// TIA Portal project "Praca_Przejsciowa_S7-1200" (V15.1)
// Vorlageprojekt für das Buch mit Zielsystem S7-1200

(* hardware
DEVICE "S7-1200-Station_1"  S7-1200 Station
   slot 0: "Baugruppenträger_0"  Rack  V1.0
   slot 1: "PLC_1"  CPU 1211C DC/DC/DC  6ES7 211-1AE40-0XB0  V4.1
DEVICE "PC-System_1"  SIMATIC PC station
   slot 0: "SIMATIC PC station"  Rail  SIMATIC PC-Station  V1.0
      slot 125: "Stationmanager"  Station_Manager  V6.0.4
   slot 1: "HMI_RT_1"  WinCC RT Advanced  6AV2 104-0xxxx-xxxx  15.1.0.0
      slot 33792: "Host interface"  Host interface
   slot 2: "IE general_1"  IE General  IE_CP  V8.2.0
*)

// ===== PLC "PLC_1"  CPU 1211C DC/DC/DC =====

VAR_GLOBAL   // PLC tag table "Standard-Variablentabelle"
   "Tag_1" AT %A0.0 : Bool;
   "Tag_2" AT %E0.0 : Bool;
   "Tag_3" AT %E0.1 : Bool;
   "Tag_4" AT %ID30 : DWord;
   "Tag_5" AT %IW32 : Word;
   "Tag_6" AT %IW36 : Int;
   "Tag_7" AT %IW40 : Int;
   "Tag_8" AT %IW30 : Int;
   "Tag_9" AT %IW3 : Word;
   "Tag_10" AT %IW34 : Int;
   "Tag_11" AT %QW30 : Int;
   "Tag_12" AT %QW32 : Int;
   "Tag_13" AT %QW34 : Int;
   "Tag_14" AT %QW40 : Int;
   "Tag_15" AT %QW42 : Int;
   "Tag_16" AT %QW44 : Int;
   "Tag_17" AT %IW38 : Int;
   "Discharge1" AT %MW10 : Int;
   "ALARM_WORD" AT %MW0 : Word;
END_VAR

// folder: DBs

DATA_BLOCK "ExchangeData"   // DB1
{ S7_Optimized_Access := 'FALSE' }
VERSION : 0.1
   VAR
      iT1_LVL : Int;   // Poziom wody w zbiorniku 1
      iT1_DIS_FL : Int;   // Przepływ na wylocie zbiornika 1
      iT1_SP : Int := 150;   // Wartość zadana regulacji w zbiorniku 1
      rT1_MV : Real;   // Wartość sterowania dla zbiornika 1
      rT1_H_REG : Real := 10.0;   // Szerokość strefy histerezy regulatora zbiornika 1
      rT1_B_REG : Real := 100.0;   // Wzmocnienie przekaźnika (Zbiornik 1)
      xT1_HH_ALM : Bool;   // Alarm poziomu HH Zbiornik 1
      xT1_H_ALM : Bool;   // Alarm poziomu H Zbiornik 1
      xT1_L_ALM : Bool;   // Alarm poziomu L Zbiornik 1
      xT1_LL_ALM : Bool;   // Alarm poziomu LL Zbiornik 1
      xT1_VLV_ALM : Bool;   // Alarm – awaria zaworu Zbiornik 1
      iT2_LVL : Int;   // Poziom wody w zbiorniku 2
      iT2_DIS_FL : Int;   // Przepływ na wylocie zbiornika 2
      iT2_SP : Int := 150;   // Wartość zadana regulacji w zbiorniku 2
      rT2_MV : Real;   // Wartość sterowania dla zbiornika 2
      rT2_P_REG : Real := 5.0;   // Wzmocnienie regulatora Zbiornik 2
      rT2_I_REG : Real := 5.0;   // Parametr I regulatora Zbiornik 2
      rT2_D_REG : Real;   // Parametr D regulatora Zbiornik 2
      xT2_HH_ALM : Bool;   // Alarm poziomu HH Zbiornik 2
      xT2_H_ALM : Bool;   // Alarm poziomu H Zbiornik 2
      xT2_L_ALM : Bool;   // Alarm poziomu L Zbiornik 2
      xT2_LL_ALM : Bool;   // Alarm poziomu LL Zbiornik 2
      xT2_VLV_ALM : Bool;   // Alarm – awaria zaworu Zbiornik 2
      iT3_LVL : Int;   // Poziom wody w zbiorniku 3
      iT3_DIS_FL : Int;   // Przepływ na wylocie zbiornika 3
      iT3_SP : Int := 150;   // Wartość zadana regulacji w zbiorniku 3
      rT3_MV : Real;   // Wartość sterowania dla zbiornika 3
      rT3_P_REG : Real := 5.0;   // Wzmocnienie regulatora Zbiornik 3
      rT3_I_REG : Real := 10.0;   // Parametr I regulatora Zbiornik 3
      rT3_B_REG : Real := 100.0;   // Wzmocnienie przekaźnika Zbiornik 3
      xT3_HH_ALM : Bool;   // Alarm poziomu HH Zbiornik 3
      xT3_H_ALM : Bool;   // Alarm poziomu H Zbiornik 3
      xT3_L_ALM : Bool;   // Alarm poziomu L Zbiornik 3
      xT3_LL_ALM : Bool;   // Alarm poziomu LL Zbiornik 3
      xT3_VLV_ALM : Bool;   // Alarm – awaria zaworu Zbiornik 3
   END_VAR
BEGIN
END_DATA_BLOCK

DATA_BLOCK "Tank1 Control_DB"   // DB4
{ S7_Optimized_Access := 'TRUE' }
VERSION : 0.1
// stored: InstanceOfName Tank1 Control
"Tank1 Control"
BEGIN
END_DATA_BLOCK

DATA_BLOCK "Disturbance Generator_DB"   // DB5
{ S7_Optimized_Access := 'TRUE' }
VERSION : 0.1
// stored: InstanceOfName Disturbance Generator
"Disturbance Generator"
BEGIN
END_DATA_BLOCK

DATA_BLOCK "Tank 2 Control_DB"   // DB8
{ S7_Optimized_Access := 'TRUE' }
VERSION : 0.1
// stored: InstanceOfName Tank 2 Control
"Tank 2 Control"
BEGIN
END_DATA_BLOCK

DATA_BLOCK "Tank 3 Control_DB"   // DB9
{ S7_Optimized_Access := 'TRUE' }
VERSION : 0.1
// stored: InstanceOfName Tank 3 Control
"Tank 3 Control"
BEGIN
END_DATA_BLOCK

// folder: IO

DATA_BLOCK "Input_DB"   // DB2
{ S7_Optimized_Access := 'TRUE' }
VERSION : 0.1
// stored: InstanceOfName Input
"Input"
BEGIN
END_DATA_BLOCK

DATA_BLOCK "Output_DB"   // DB3
{ S7_Optimized_Access := 'TRUE' }
VERSION : 0.1
// stored: InstanceOfName Output
"Output"
BEGIN
END_DATA_BLOCK

// folder: (top level)

FUNCTION_BLOCK "Tank1 Control"   // FB3, LAD
{ S7_Optimized_Access := 'TRUE' }
VERSION : 0.1
   VAR_INPUT
      Level : Int;
      SP : Int := 150;
      h_reg : Real := 10.0;
      B_reg : Real := 100.0;
      HH_LVL : Int := 280;
      H_LVL : Int := 250;
      L_LVL : Int := 50;
      LL_LVL : Int := 20;
   END_VAR
   VAR_OUTPUT
      HH_Alarm : Bool;
      H_Alarm : Bool;
      L_Alarm : Bool;
      LL_Alarm : Bool;
      Vlv_Pos_Alarm : Bool;
      MV : Real;
   END_VAR
   VAR
      prev_control : Bool;
      control_action : Bool;
   END_VAR
BEGIN

REGION Network 1 (SCL)
   REGION Level control

       IF #Level < #SP - #h_reg THEN
           #control_action := 1;
       ELSIF #Level > #SP + #h_reg THEN
           #control_action := 0;
       ELSE
           #control_action := #prev_control;
       END_IF;

       #prev_control := #control_action;

       #MV := BOOL_TO_INT(#control_action) * #B_reg;


   END_REGION


   REGION ALARMS
       #HH_Alarm := FALSE;
       #H_Alarm := FALSE;
       #LL_Alarm := FALSE;
       #L_Alarm := FALSE;

       IF #Level > #HH_LVL THEN
           #HH_Alarm := TRUE;
       ELSIF #Level > #H_LVL THEN
           #H_Alarm := TRUE;
       END_IF;

       IF #Level < #LL_LVL THEN
           #LL_Alarm := TRUE;
       ELSIF #Level < #L_LVL THEN
           #L_Alarm := TRUE;
       END_IF;

   END_REGION
END_REGION
END_FUNCTION_BLOCK

FUNCTION_BLOCK "Disturbance Generator"   // FB4, LAD
{ S7_Optimized_Access := 'TRUE' }
VERSION : 0.1
   VAR_INPUT
      minOpen : Int;
      maxOpen : Int := 100;
   END_VAR
   VAR_OUTPUT
      iT1_Dis_vlv : Int;
      iT2_Dis_vlv : Int;
      iT3_Dis_vlv : Int;
   END_VAR
   VAR
      rDistrbance_T1 : Real := 50.0;
      rDistrbance_T2 : Real := 50.0;
      rDistrbance_T3 : Real := 50.0;
      rDisturbanceDesire : Real := 40.0;
      xDistrubanceRising : Bool;
   END_VAR
   VAR_TEMP
      temp_time : DTL;
      Seed1 : Real;
      Seed2 : Real;
      dist1 : Real;
      dist2 : Real;
      dist3 : Real;
   END_VAR
BEGIN

REGION Network 1 (SCL)
   // Symulacja zmian otwarcia zaworu na wyjściu jako zakłócenia
   // Seed generation from system clock
   #Seed1 := RD_SYS_T(#temp_time);
   #Seed1 := #temp_time.SECOND;
   #Seed2 := #temp_time.NANOSECOND;
   //fast and randomly changing distrubance
   #dist1 := SIN(#Seed1) + SIN(#Seed2);
   #dist1 := COS(#Seed1) + SIN(#Seed2);
   #dist1 := COS(#Seed1) + COS(#Seed2);

   // Slowly changing opennig between 20-70%
   IF #xDistrubanceRising THEN
       #rDisturbanceDesire := #rDisturbanceDesire + 0.05;
   ELSE
       #rDisturbanceDesire := #rDisturbanceDesire - 0.05;
   END_IF;

   IF #rDisturbanceDesire < 20.0 THEN
       #xDistrubanceRising := TRUE;
   ELSIF #rDisturbanceDesire > 70.0 THEN
       #xDistrubanceRising := FALSE;
   END_IF;

   // Position is sum of random distrubance and factor pushing it to
   // slowly changing desired position
   #rDistrbance_T1 := #rDistrbance_T1 + 0.1 * #dist1 + 0.01*(#rDisturbanceDesire - #rDistrbance_T1);
   #rDistrbance_T2 := #rDistrbance_T2 + 0.1 * #dist2 + 0.01 * (#rDisturbanceDesire - #rDistrbance_T2);
   #rDistrbance_T3 := #rDistrbance_T3 + 0.1 * #dist3 + 0.01 * (#rDisturbanceDesire - #rDistrbance_T3);

   // Position limited between 5-95%
   #iT1_Dis_vlv := LIMIT(MN := 5, IN := #rDistrbance_T1, MX := 95);
   #iT2_Dis_vlv := LIMIT(MN := 5, IN := #rDistrbance_T2, MX := 95);
   #iT3_Dis_vlv := LIMIT(MN := 5, IN := #rDistrbance_T3, MX := 95);
END_REGION
END_FUNCTION_BLOCK

FUNCTION_BLOCK "Tank 2 Control"   // FB5, SCL
{ S7_Optimized_Access := 'TRUE' }
VERSION : 0.1
   VAR_INPUT
      Level : Int := 0;
      SP : Int := 150;
      P_reg : Real := 10.0;
      I_reg : Real := 10.0;
      HH_LVL : Int := 280;
      H_LVL : Int := 250;
      L_LVL : Int := 50;
      LL_LVL : Int := 20;
   END_VAR
   VAR_OUTPUT
      HH_Alarm : Bool := false;
      H_Alarm : Bool := false;
      L_Alarm : Bool := false;
      LL_Alarm : Bool := false;
      Vlv_Pos_Alarm : Bool := false;
      MV : Real := 0.0;
   END_VAR
   VAR
      I_action : Real := 0.0;
      Error : Real;
      Executed : Bool;
   END_VAR
   VAR_TEMP
      P_action : Real;
   END_VAR
   VAR CONSTANT
      Interval : Time := T#100ms;
      rInterval_ms : Real := 100.0;
   END_VAR
BEGIN
   // PID opration handled by OB30
   // for constant interval time

   REGION ALARMS
       #HH_Alarm := FALSE;
       #H_Alarm := FALSE;
       #LL_Alarm := FALSE;
       #L_Alarm := FALSE;

       IF #Level > #HH_LVL THEN
           #HH_Alarm := TRUE;
       ELSIF #Level > #H_LVL THEN
           #H_Alarm := TRUE;
       END_IF;

       IF #Level < #LL_LVL THEN
           #LL_Alarm := TRUE;
       ELSIF #Level < #L_LVL THEN
           #L_Alarm := TRUE;
       END_IF;

   END_REGION
END_FUNCTION_BLOCK

FUNCTION_BLOCK "Tank 3 Control"   // FB6, LAD
{ S7_Optimized_Access := 'TRUE' }
VERSION : 0.1
   VAR_INPUT
      Level : Int;
      SP : Int := 150;
      P_reg : Real := 5.0;
      I_reg : Real := 10.0;
      B_reg : Real := 100.0;
      HH_LVL : Int := 280;
      H_LVL : Int := 250;
      L_LVL : Int := 50;
      LL_LVL : Int := 20;
   END_VAR
   VAR_OUTPUT
      HH_Alarm : Bool := false;
      H_Alarm : Bool := false;
      L_Alarm : Bool := false;
      LL_Alarm : Bool := false;
      Vlv_Pos_Alarm : Bool := false;
      MV : Real := 0.0;
   END_VAR
   VAR
      I_action : Real := 0.0;
      Error : Real := 0.0;
      Ref_sig : Real := 0.0;
      Control_sig : Real := 0.0;
      Ref_sig_period : Real := 5.0;   // okres sygnały piłokształtnego
   END_VAR
BEGIN

REGION Network 1
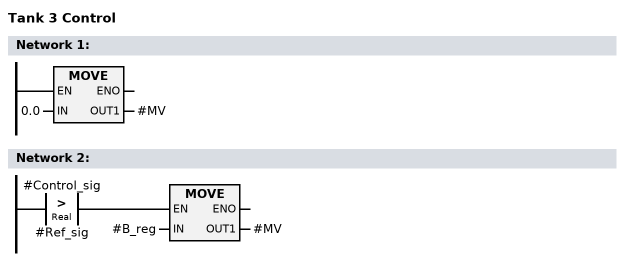
   RUNG wire#powerrail
      Move(in := 0.0, out1 => #MV)
   END_RUNG
   // the same network as SCL:
   #MV := 0.0;
END_REGION

REGION Network 2
   RUNG wire#powerrail
      { S7_Templates := "SrcType := Real" } GT_Contact(in1 := #Control_sig, in2 := #Ref_sig)
      Move(in := #B_reg, out1 => #MV)
   END_RUNG
   // the same network as SCL:
   IF #Control_sig > #Ref_sig THEN #MV := #B_reg; END_IF;
END_REGION

REGION Network 3 (SCL)
   // PID opration handled by OB31
   // for constant interval time

   REGION ALARMS
       #HH_Alarm := FALSE;
       #H_Alarm := FALSE;
       #LL_Alarm := FALSE;
       #L_Alarm := FALSE;

       IF #Level > #HH_LVL THEN
           #HH_Alarm := TRUE;
       ELSIF #Level > #H_LVL THEN
           #H_Alarm := TRUE;
       END_IF;

       IF #Level < #LL_LVL THEN
           #LL_Alarm := TRUE;
       ELSIF #Level < #L_LVL THEN
           #L_Alarm := TRUE;
       END_IF;

   END_REGION
END_REGION
END_FUNCTION_BLOCK

ORGANIZATION_BLOCK "Main"   // OB1, LAD, ProgramCycle
TITLE = "Main Program Sweep (Cycle)"
{ S7_Optimized_Access := 'TRUE' }
VERSION : 0.1
   VAR_INPUT
      Initial_Call : Bool;   // Initial call of this OB
      Remanence : Bool;   // =True, if remanent data are available
   END_VAR
BEGIN

REGION Network 1: Konnektierungsbaustein für PLC-Lab
   // Im Netzwerk 1 wird der Konnektierungsbaustein für PLC-Lab aufgerufen.
   // Dieser Aufruf darf nicht entfernt werden!
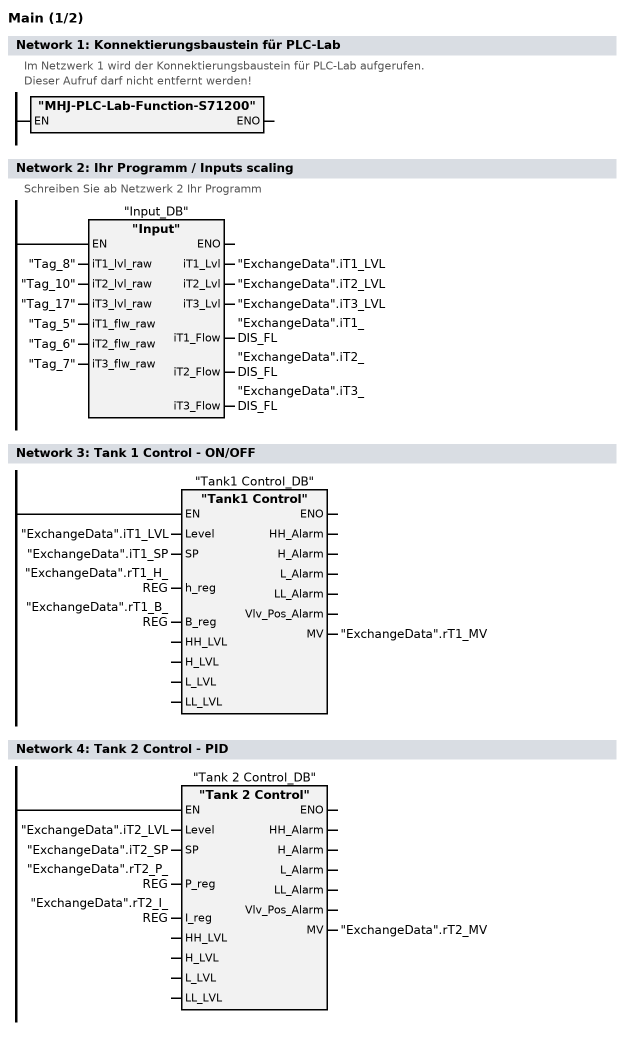
   RUNG wire#powerrail
      "MHJ-PLC-Lab-Function-S71200"()
   END_RUNG
   // the same network as SCL:
   "MHJ-PLC-Lab-Function-S71200"();
END_REGION

REGION Network 2: Ihr Programm / Inputs scaling
   // Schreiben Sie ab Netzwerk 2 Ihr Programm
   RUNG wire#powerrail
      "Input_DB"(iT1_lvl_raw := "Tag_8", iT2_lvl_raw := "Tag_10", iT3_lvl_raw := "Tag_17", iT1_flw_raw := "Tag_5", iT2_flw_raw := "Tag_6", iT3_flw_raw := "Tag_7", iT1_Lvl => "ExchangeData".iT1_LVL, iT2_Lvl => "ExchangeData".iT2_LVL, iT3_Lvl => "ExchangeData".iT3_LVL, iT1_Flow => "ExchangeData".iT1_DIS_FL, iT2_Flow => "ExchangeData".iT2_DIS_FL, iT3_Flow => "ExchangeData".iT3_DIS_FL)
   END_RUNG
   // the same network as SCL:
   "Input_DB"(iT1_lvl_raw := "Tag_8",   // "Input"
              iT2_lvl_raw := "Tag_10",
              iT3_lvl_raw := "Tag_17",
              iT1_flw_raw := "Tag_5",
              iT2_flw_raw := "Tag_6",
              iT3_flw_raw := "Tag_7",
              iT1_Lvl => "ExchangeData".iT1_LVL,
              iT2_Lvl => "ExchangeData".iT2_LVL,
              iT3_Lvl => "ExchangeData".iT3_LVL,
              iT1_Flow => "ExchangeData".iT1_DIS_FL,
              iT2_Flow => "ExchangeData".iT2_DIS_FL,
              iT3_Flow => "ExchangeData".iT3_DIS_FL);
END_REGION

REGION Network 3: Tank 1 Control - ON/OFF
   RUNG wire#powerrail
      "Tank1 Control_DB"(Level := "ExchangeData".iT1_LVL, SP := "ExchangeData".iT1_SP, h_reg := "ExchangeData".rT1_H_REG, B_reg := "ExchangeData".rT1_B_REG, HH_LVL :=, H_LVL :=, L_LVL :=, LL_LVL :=, HH_Alarm =>, H_Alarm =>, L_Alarm =>, LL_Alarm =>, Vlv_Pos_Alarm =>, MV => "ExchangeData".rT1_MV)
   END_RUNG
   // the same network as SCL:
   "Tank1 Control_DB"(Level := "ExchangeData".iT1_LVL,   // "Tank1 Control"
                      SP := "ExchangeData".iT1_SP,
                      h_reg := "ExchangeData".rT1_H_REG,
                      B_reg := "ExchangeData".rT1_B_REG,
                      MV => "ExchangeData".rT1_MV);
END_REGION

REGION Network 4: Tank 2 Control - PID
   RUNG wire#powerrail
      "Tank 2 Control_DB"(Level := "ExchangeData".iT2_LVL, SP := "ExchangeData".iT2_SP, P_reg := "ExchangeData".rT2_P_REG, I_reg := "ExchangeData".rT2_I_REG, HH_LVL :=, H_LVL :=, L_LVL :=, LL_LVL :=, HH_Alarm =>, H_Alarm =>, L_Alarm =>, LL_Alarm =>, Vlv_Pos_Alarm =>, MV => "ExchangeData".rT2_MV)
   END_RUNG
   // the same network as SCL:
   "Tank 2 Control_DB"(Level := "ExchangeData".iT2_LVL,   // "Tank 2 Control"
                       SP := "ExchangeData".iT2_SP,
                       P_reg := "ExchangeData".rT2_P_REG,
                       I_reg := "ExchangeData".rT2_I_REG,
                       MV => "ExchangeData".rT2_MV);
END_REGION

REGION Network 5: Tank 3 Control - PID PWM
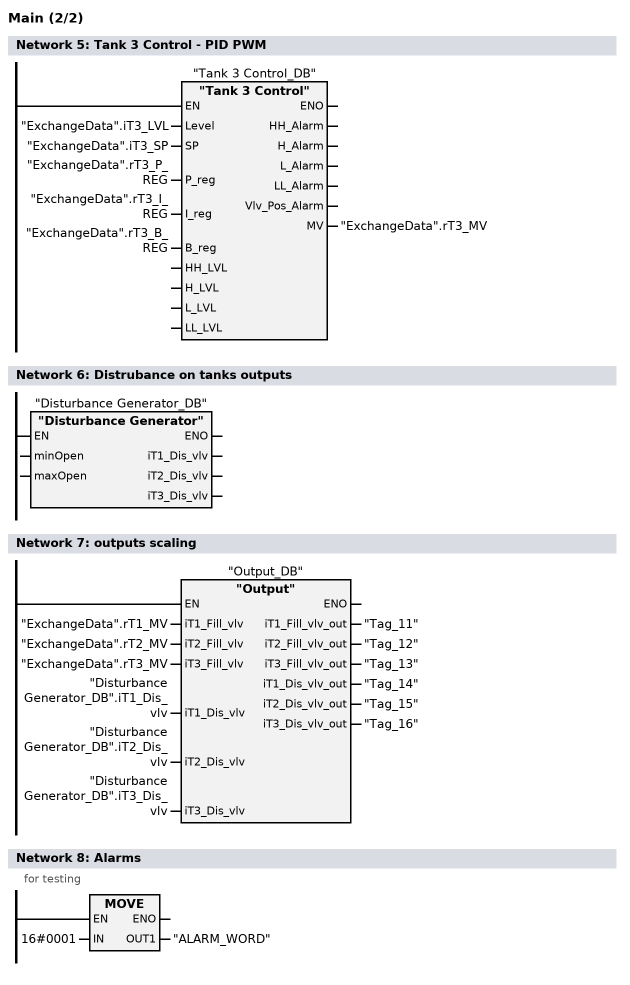
   RUNG wire#powerrail
      "Tank 3 Control_DB"(Level := "ExchangeData".iT3_LVL, SP := "ExchangeData".iT3_SP, P_reg := "ExchangeData".rT3_P_REG, I_reg := "ExchangeData".rT3_I_REG, B_reg := "ExchangeData".rT3_B_REG, HH_LVL :=, H_LVL :=, L_LVL :=, LL_LVL :=, HH_Alarm =>, H_Alarm =>, L_Alarm =>, LL_Alarm =>, Vlv_Pos_Alarm =>, MV => "ExchangeData".rT3_MV)
   END_RUNG
   // the same network as SCL:
   "Tank 3 Control_DB"(Level := "ExchangeData".iT3_LVL,   // "Tank 3 Control"
                       SP := "ExchangeData".iT3_SP,
                       P_reg := "ExchangeData".rT3_P_REG,
                       I_reg := "ExchangeData".rT3_I_REG,
                       B_reg := "ExchangeData".rT3_B_REG,
                       MV => "ExchangeData".rT3_MV);
END_REGION

REGION Network 6: Distrubance on tanks outputs
   RUNG wire#powerrail
      "Disturbance Generator_DB"(minOpen :=, maxOpen :=, iT1_Dis_vlv =>, iT2_Dis_vlv =>, iT3_Dis_vlv =>)
   END_RUNG
   // the same network as SCL:
   "Disturbance Generator_DB"();   // "Disturbance Generator"
END_REGION

REGION Network 7: outputs scaling
   RUNG wire#powerrail
      "Output_DB"(iT1_Fill_vlv := "ExchangeData".rT1_MV, iT2_Fill_vlv := "ExchangeData".rT2_MV, iT3_Fill_vlv := "ExchangeData".rT3_MV, iT1_Dis_vlv := "Disturbance Generator_DB".iT1_Dis_vlv, iT2_Dis_vlv := "Disturbance Generator_DB".iT2_Dis_vlv, iT3_Dis_vlv := "Disturbance Generator_DB".iT3_Dis_vlv, iT1_Fill_vlv_out => "Tag_11", iT2_Fill_vlv_out => "Tag_12", iT3_Fill_vlv_out => "Tag_13", iT1_Dis_vlv_out => "Tag_14", iT2_Dis_vlv_out => "Tag_15", iT3_Dis_vlv_out => "Tag_16")
   END_RUNG
   // the same network as SCL:
   "Output_DB"(iT1_Fill_vlv := "ExchangeData".rT1_MV,   // "Output"
               iT2_Fill_vlv := "ExchangeData".rT2_MV,
               iT3_Fill_vlv := "ExchangeData".rT3_MV,
               iT1_Dis_vlv := "Disturbance Generator_DB".iT1_Dis_vlv,
               iT2_Dis_vlv := "Disturbance Generator_DB".iT2_Dis_vlv,
               iT3_Dis_vlv := "Disturbance Generator_DB".iT3_Dis_vlv,
               iT1_Fill_vlv_out => "Tag_11",
               iT2_Fill_vlv_out => "Tag_12",
               iT3_Fill_vlv_out => "Tag_13",
               iT1_Dis_vlv_out => "Tag_14",
               iT2_Dis_vlv_out => "Tag_15",
               iT3_Dis_vlv_out => "Tag_16");
END_REGION

REGION Network 8: Alarms
   // for testing
   RUNG wire#powerrail
      Move(in := 16#0001, out1 => "ALARM_WORD")
   END_RUNG
   // the same network as SCL:
   "ALARM_WORD" := 16#0001;
END_REGION
END_ORGANIZATION_BLOCK

ORGANIZATION_BLOCK "PID_2"   // OB30, LAD, CyclicInterrupt
{ S7_Optimized_Access := 'TRUE' }
VERSION : 0.1
   VAR_INPUT
      Initial_Call : Bool;   // Initial call of this OB
      Event_Count : Int;   // Events discarded
   END_VAR
   VAR_TEMP
      Error : Real;
      P_action : Real;
      I_action : Real;
   END_VAR
BEGIN

REGION Network 1 (SCL)
   #Error :="Tank 2 Control_DB".SP -"Tank 2 Control_DB".Level;

   #P_action := #Error * "Tank 2 Control_DB".P_reg;

   IF "Tank 2 Control_DB".MV < 100.0 AND "Tank 2 Control_DB".MV > 0.0 THEN
       "Tank 2 Control_DB".I_action := "Tank 2 Control_DB".I_action + "Tank 2 Control_DB".P_reg * (#Error / "Tank 2 Control_DB".I_reg * 0.1);
   END_IF;

   "Tank 2 Control_DB".MV := #P_action + "Tank 2 Control_DB".I_action;
   "Tank 2 Control_DB".MV := LIMIT(MN := 0.0, IN := "Tank 2 Control_DB".MV, MX := 100.0);
END_REGION
END_ORGANIZATION_BLOCK

ORGANIZATION_BLOCK "PID_3"   // OB31, SCL, CyclicInterrupt
{ S7_Optimized_Access := 'TRUE' }
VERSION : 0.1
   VAR_INPUT
      Initial_Call : Bool;   // Initial call of this OB
      Event_Count : Int;   // Events discarded
   END_VAR
   VAR_TEMP
      Error : Real;
      P_action : Real;
      I_action : Real;
      Ref_sig_increment : Real;
   END_VAR
BEGIN
   #Error := "Tank 3 Control_DB".SP - "Tank 3 Control_DB".Level;

   #P_action := #Error * "Tank 3 Control_DB".P_reg;

   IF "Tank 3 Control_DB".Control_sig < 100.0 AND "Tank 3 Control_DB".Control_sig > 0.0 THEN
       "Tank 3 Control_DB".I_action := "Tank 3 Control_DB".I_action + "Tank 3 Control_DB".P_reg * (#Error / "Tank 3 Control_DB".I_reg * 0.1);
   END_IF;

   "Tank 3 Control_DB".Control_sig := #P_action + "Tank 3 Control_DB".I_action;
   "Tank 3 Control_DB".Control_sig := LIMIT(MN := 0.0, IN := "Tank 3 Control_DB".Control_sig, MX := 100.0);

   // Reference signal conditioning
   #Ref_sig_increment := 100.0 / 10.0 / "Tank 3 Control_DB".Ref_sig_period;
   "Tank 3 Control_DB".Ref_sig := "Tank 3 Control_DB".Ref_sig + #Ref_sig_increment;

   IF "Tank 3 Control_DB".Ref_sig > 100.0 THEN
       "Tank 3 Control_DB".Ref_sig := 0;
   END_IF;
END_ORGANIZATION_BLOCK

// folder: IO

FUNCTION_BLOCK "Input"   // FB1, LAD
{ S7_Optimized_Access := 'TRUE' }
VERSION : 0.1
   VAR_INPUT
      iT1_lvl_raw : Int;
      iT2_lvl_raw : Int;
      iT3_lvl_raw : Int;
      iT1_flw_raw : Int;
      iT2_flw_raw : Int;
      iT3_flw_raw : Int;
   END_VAR
   VAR_OUTPUT
      iT1_Lvl : Int;
      iT2_Lvl : Int;
      iT3_Lvl : Int;
      iT1_Flow : Int;
      iT2_Flow : Int;
      iT3_Flow : Int;
   END_VAR
BEGIN

REGION Network 1
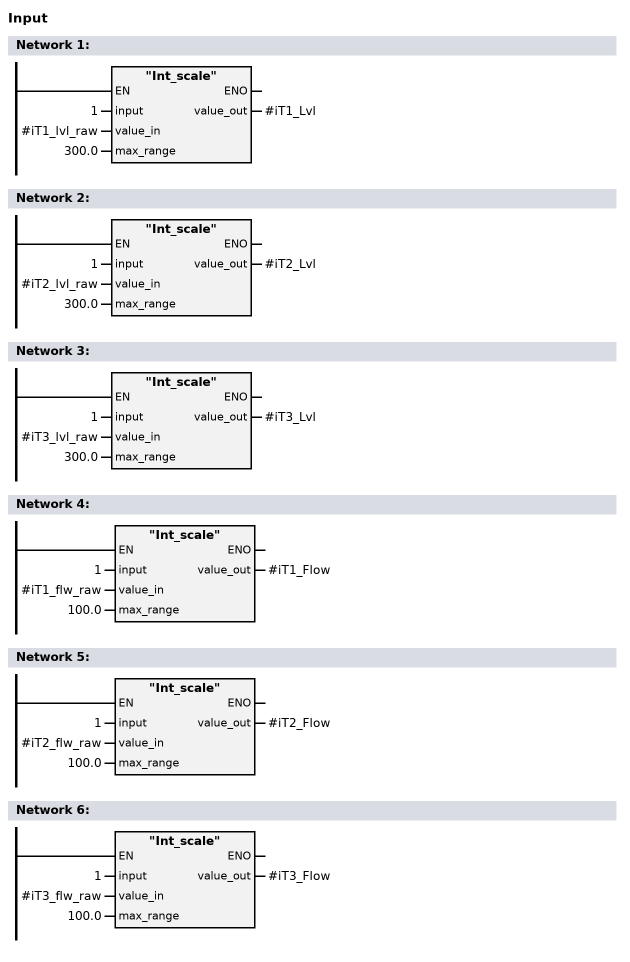
   RUNG wire#powerrail
      "Int_scale"(input := 1, value_in := #iT1_lvl_raw, max_range := 300.0, value_out => #iT1_Lvl)
   END_RUNG
   // the same network as SCL:
   "Int_scale"(input := 1, value_in := #iT1_lvl_raw, max_range := 300.0, value_out => #iT1_Lvl);
END_REGION

REGION Network 2
   RUNG wire#powerrail
      "Int_scale"(input := 1, value_in := #iT2_lvl_raw, max_range := 300.0, value_out => #iT2_Lvl)
   END_RUNG
   // the same network as SCL:
   "Int_scale"(input := 1, value_in := #iT2_lvl_raw, max_range := 300.0, value_out => #iT2_Lvl);
END_REGION

REGION Network 3
   RUNG wire#powerrail
      "Int_scale"(input := 1, value_in := #iT3_lvl_raw, max_range := 300.0, value_out => #iT3_Lvl)
   END_RUNG
   // the same network as SCL:
   "Int_scale"(input := 1, value_in := #iT3_lvl_raw, max_range := 300.0, value_out => #iT3_Lvl);
END_REGION

REGION Network 4
   RUNG wire#powerrail
      "Int_scale"(input := 1, value_in := #iT1_flw_raw, max_range := 100.0, value_out => #iT1_Flow)
   END_RUNG
   // the same network as SCL:
   "Int_scale"(input := 1, value_in := #iT1_flw_raw, max_range := 100.0, value_out => #iT1_Flow);
END_REGION

REGION Network 5
   RUNG wire#powerrail
      "Int_scale"(input := 1, value_in := #iT2_flw_raw, max_range := 100.0, value_out => #iT2_Flow)
   END_RUNG
   // the same network as SCL:
   "Int_scale"(input := 1, value_in := #iT2_flw_raw, max_range := 100.0, value_out => #iT2_Flow);
END_REGION

REGION Network 6
   RUNG wire#powerrail
      "Int_scale"(input := 1, value_in := #iT3_flw_raw, max_range := 100.0, value_out => #iT3_Flow)
   END_RUNG
   // the same network as SCL:
   "Int_scale"(input := 1, value_in := #iT3_flw_raw, max_range := 100.0, value_out => #iT3_Flow);
END_REGION
END_FUNCTION_BLOCK

FUNCTION_BLOCK "Output"   // FB2, LAD
{ S7_Optimized_Access := 'TRUE' }
VERSION : 0.1
   VAR_INPUT
      iT1_Fill_vlv : Int;
      iT2_Fill_vlv : Int;
      iT3_Fill_vlv : Int;
      iT1_Dis_vlv : Int;
      iT2_Dis_vlv : Int;
      iT3_Dis_vlv : Int;
   END_VAR
   VAR_OUTPUT
      iT1_Fill_vlv_out : Int;
      iT2_Fill_vlv_out : Int;
      iT3_Fill_vlv_out : Int;
      iT1_Dis_vlv_out : Int;
      iT2_Dis_vlv_out : Int;
      iT3_Dis_vlv_out : Int;
   END_VAR
BEGIN

REGION Network 1
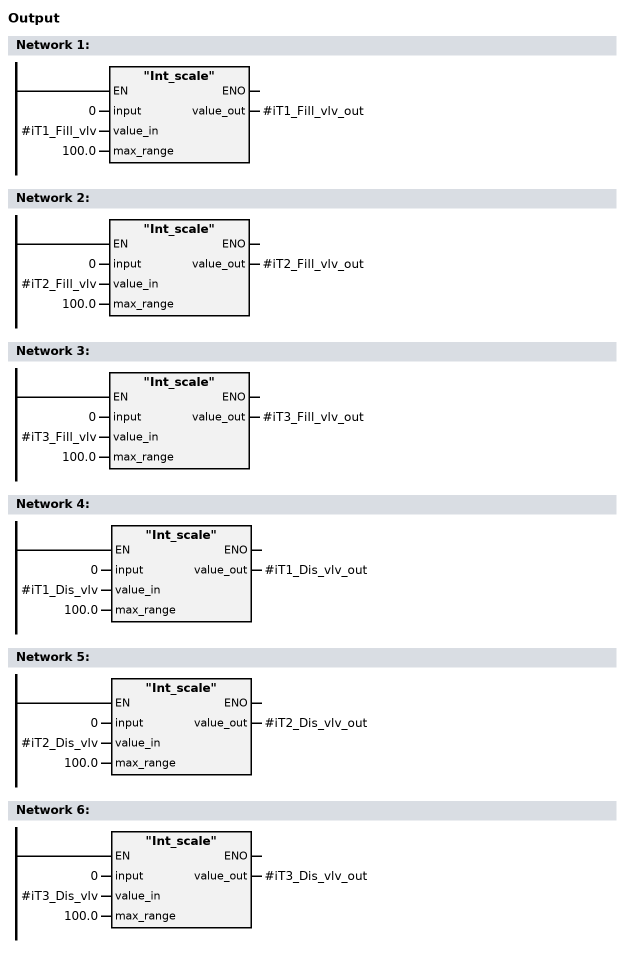
   RUNG wire#powerrail
      "Int_scale"(input := 0, value_in := #iT1_Fill_vlv, max_range := 100.0, value_out => #iT1_Fill_vlv_out)
   END_RUNG
   // the same network as SCL:
   "Int_scale"(input := 0, value_in := #iT1_Fill_vlv, max_range := 100.0, value_out => #iT1_Fill_vlv_out);
END_REGION

REGION Network 2
   RUNG wire#powerrail
      "Int_scale"(input := 0, value_in := #iT2_Fill_vlv, max_range := 100.0, value_out => #iT2_Fill_vlv_out)
   END_RUNG
   // the same network as SCL:
   "Int_scale"(input := 0, value_in := #iT2_Fill_vlv, max_range := 100.0, value_out => #iT2_Fill_vlv_out);
END_REGION

REGION Network 3
   RUNG wire#powerrail
      "Int_scale"(input := 0, value_in := #iT3_Fill_vlv, max_range := 100.0, value_out => #iT3_Fill_vlv_out)
   END_RUNG
   // the same network as SCL:
   "Int_scale"(input := 0, value_in := #iT3_Fill_vlv, max_range := 100.0, value_out => #iT3_Fill_vlv_out);
END_REGION

REGION Network 4
   RUNG wire#powerrail
      "Int_scale"(input := 0, value_in := #iT1_Dis_vlv, max_range := 100.0, value_out => #iT1_Dis_vlv_out)
   END_RUNG
   // the same network as SCL:
   "Int_scale"(input := 0, value_in := #iT1_Dis_vlv, max_range := 100.0, value_out => #iT1_Dis_vlv_out);
END_REGION

REGION Network 5
   RUNG wire#powerrail
      "Int_scale"(input := 0, value_in := #iT2_Dis_vlv, max_range := 100.0, value_out => #iT2_Dis_vlv_out)
   END_RUNG
   // the same network as SCL:
   "Int_scale"(input := 0, value_in := #iT2_Dis_vlv, max_range := 100.0, value_out => #iT2_Dis_vlv_out);
END_REGION

REGION Network 6
   RUNG wire#powerrail
      "Int_scale"(input := 0, value_in := #iT3_Dis_vlv, max_range := 100.0, value_out => #iT3_Dis_vlv_out)
   END_RUNG
   // the same network as SCL:
   "Int_scale"(input := 0, value_in := #iT3_Dis_vlv, max_range := 100.0, value_out => #iT3_Dis_vlv_out);
END_REGION
END_FUNCTION_BLOCK

FUNCTION "Int_scale" : Void   // FC1, SCL
{ S7_Optimized_Access := 'TRUE' }
VERSION : 0.1
   VAR_INPUT
      input : Bool;
      value_in : Int;
      max_range : Real;
   END_VAR
   VAR_OUTPUT
      value_out : Int;
   END_VAR
   VAR_TEMP
      scale_unit : Real;
   END_VAR
   VAR CONSTANT
      Int_range : Int := 27648;
   END_VAR
BEGIN
   IF #input = 1 THEN
       #scale_unit := INT_TO_REAL(#value_in) / INT_TO_REAL(#Int_range);
       #value_out := REAL_TO_INT(#scale_unit * #max_range);
   END_IF;

   IF #input = 0 THEN
       #scale_unit := INT_TO_REAL(#value_in)/#max_range;
       #value_out := REAL_TO_INT(#scale_unit *#Int_range);
   END_IF;
END_FUNCTION

FUNCTION "MHJ-PLC-Lab-Function-S71200" : Void   // FC9000, SCL
{ S7_Optimized_Access := 'TRUE' }
VERSION : 0.1
   VAR_TEMP
      rdTimeReturn : Int;
      outputTime : DTL;
      SyncVal : Byte;
      forVal : Int;
      forVal_2 : Int;
      Value : Byte;
   END_VAR
   VAR CONSTANT
      CompVal : Byte := 16#34;
      Value_01 : Byte := 16#11;
      Value_01_DW : DWord := 16#A165_D992;
      Value_02_DW : DWord := 16#58BE_4401;
   END_VAR
BEGIN

   #Value:=PEEK(area := 16#82,
        dbNumber := 0,
        byteOffset := 511);
   #Value := #Value + 1;

   POKE(area := 16#82,
        dbNumber := 0,
        byteOffset := 511,
        value := #Value);

   POKE(area:=16#81,
        dbNumber:=0,
        byteOffset:=1016,
        value:=#Value_01_DW);
   POKE(area := 16#81,
        dbNumber := 0,
        byteOffset := 1020,
        value := #Value_02_DW);

   POKE(area := 16#81,
        dbNumber := 0,
        byteOffset := 511,
        value := B#16#00);

   FOR #forVal := 0 TO 120 DO
       FOR #forVal_2:=0 TO 10 DO
           #rdTimeReturn:=RD_SYS_T(#outputTime);
           #rdTimeReturn := WR_SYS_T(#outputTime);
           #rdTimeReturn := RD_SYS_T(#outputTime);
           #rdTimeReturn := WR_SYS_T(#outputTime);
       END_FOR;
       #SyncVal:= PEEK(area := 16#81,
                      dbNumber := 0,
                      byteOffset := 511);
       IF #SyncVal = #CompVal THEN
          GOTO M_1;
       END_IF;
   END_FOR;
   RETURN;

   M_1:
   POKE(area := 16#81,
        dbNumber := 0,
        byteOffset := 511,
        value := B#16#0);
END_FUNCTION

(* ===== HMI "HMI_RT_1" =====
system functions are stored by id; their names below are inferred from use
connection "Connection_1": ETHERNET, S7_1200_OMS
connection "HMI_Connection_1": ETHERNET, S7_1200_OMS

HMI tags "Default tag table"
   "T1_LVL" : Int = PLC ExchangeData.iT1_LVL AT %DB1.DBW0, 1 s
   "T1_MV" : Real = PLC ExchangeData.rT1_MV AT %DB1.DBD6, 1 s
   "T1_Dis_fl" : Int = PLC ExchangeData.iT1_DIS_FL AT %DB1.DBW2, 1 s
   "T1_Dis" : Int = PLC "Disturbance Generator_DB".iT1_Dis_vlv AT %MW10, 1 s
   "T1_SP" : Int = PLC ExchangeData.iT1_SP AT %DB1.DBW4, 1 s
   "T1_H_reg" : Real = PLC ExchangeData.rT1_H_REG AT %DB1.DBD10, 1 s
   "T1_B_reg" : Real = PLC ExchangeData.rT1_B_REG AT %DB1.DBD14, 1 s
   "T2_Dis_fl" : Int = PLC ExchangeData.iT2_DIS_FL AT %DB1.DBW22, 1 s
   "T2_Dis" : Int = PLC "Disturbance Generator_DB".iT2_Dis_vlv AT %DB1.DBW0, 1 s
   "T2_MV" : Real = PLC ExchangeData.rT2_MV AT %DB1.DBD26, 1 s
   "T2_LVL" : Int = PLC ExchangeData.iT2_LVL AT %DB1.DBW20, 1 s
   "T2_SP" : Int = PLC ExchangeData.iT2_SP AT %DB1.DBW24, 1 s
   "T2_P_reg" : Real = PLC ExchangeData.rT2_P_REG AT %DB1.DBD30, 1 s
   "T2_I_reg" : Real = PLC ExchangeData.rT2_I_REG AT %DB1.DBD34, 1 s
   "T3_I_reg" : Real = PLC ExchangeData.rT3_I_REG AT %DB1.DBD58, 1 s
   "T3_P_reg" : Real = PLC ExchangeData.rT3_P_REG AT %DB1.DBD54, 1 s
   "T3_LVL" : Int = PLC ExchangeData.iT3_LVL AT %DB1.DBW44, 1 s
   "T3_Ref" : Real = PLC "Tank 3 Control_DB".Ref_sig AT %DB1.DBD0, 1 s
   "T3_MV" : Real = PLC ExchangeData.rT3_MV AT %DB1.DBD50, 1 s
   "T3_Dis" : Int = PLC "Disturbance Generator_DB".iT3_Dis_vlv AT %DB1.DBW0, 1 s
   "T3_SP" : Int = PLC ExchangeData.iT3_SP AT %DB1.DBW48, 1 s
   "T3_PID_CTRL" : Real = PLC "Tank 3 Control_DB".Control_sig AT %DB1.DBW0, 1 s
   "T3_Dis_fl" : Int = PLC ExchangeData.iT3_DIS_FL AT %DB1.DBW46, 1 s
   "T3_B_reg" : Real = PLC ExchangeData.rT3_B_REG AT %DB1.DBD62, 1 s

HMI tags "Alarms"
   "T1_LL" : Bool = PLC ExchangeData.xT1_LL_ALM AT %DB1.DBX18.3, 1 s
   "T1_L" : Bool = PLC ExchangeData.xT1_L_ALM AT %DB1.DBX18.2, 1 s
   "T1_H" : Bool = PLC ExchangeData.xT1_H_ALM AT %DB1.DBX18.1, 1 s
   "T1_HH" : Bool = PLC ExchangeData.xT1_HH_ALM AT %DB1.DBX18.0, 1 s
   "T2_LL" : Bool = PLC ExchangeData.xT2_LL_ALM AT %DB1.DBX42.3, 1 s
   "T2_L" : Bool = PLC ExchangeData.xT2_L_ALM AT %DB1.DBX42.2, 1 s
   "T2_H" : Bool = PLC ExchangeData.xT2_H_ALM AT %DB1.DBX42.1, 1 s
   "T2_HH" : Bool = PLC ExchangeData.xT2_HH_ALM AT %DB1.DBX42.0, 1 s
   "T3_LL" : Bool = PLC ExchangeData.xT3_LL_ALM AT %DB1.DBX66.3, 1 s
   "T3_L" : Bool = PLC ExchangeData.xT3_L_ALM AT %DB1.DBX66.2, 1 s
   "T3_H" : Bool = PLC ExchangeData.xT3_H_ALM AT %DB1.DBX66.1, 1 s
   "T3_HH" : Bool = PLC ExchangeData.xT3_HH_ALM AT %DB1.DBX66.0, 1 s
   "T1_vlv_alm" : Bool = PLC ExchangeData.xT1_VLV_ALM AT %DB1.DBX18.4, 1 s
   "T2_vlv_alm" : Bool = PLC ExchangeData.xT2_VLV_ALM AT %DB1.DBX42.4, 1 s
   "ALARMS" : Word = PLC ALARM_WORD AT %MW0, 1 s
   "Acknowledge" : Int AT %DB1.DBX0.0

discrete alarms
   1: 'Tank1 Level LL', class Errors, trigger "ALARMS" bit 0
   2: 'Tank1 Level L', class Warnings, trigger "ALARMS" bit 1
   3: 'Tank1 Level H', class Warnings, trigger "ALARMS" bit 2
   4: 'Tank1 Level HH', class Errors, trigger "ALARMS" bit 3
   5: 'Tank2 Level LL', class Errors, trigger "ALARMS" bit 4
   6: 'Tank2 Level L', class Warnings, trigger "ALARMS" bit 5
   7: 'Tank2 Level H', class Warnings, trigger "ALARMS" bit 6
   8: 'Tank2 Level HH', class Errors, trigger "ALARMS" bit 7
   9: 'Tank3 Level LL', class Errors, trigger "ALARMS" bit 8
   11: 'Tank3 Level H', class Warnings, trigger "ALARMS" bit 10
   12: 'Tank3 Level HH', class Errors, trigger "ALARMS" bit 11
   13: 'Tank1 Valve Error', class Errors, trigger "ALARMS" bit 12
   14: 'Tank2 Valve Error', class Errors, trigger "ALARMS" bit 13
   15: 'Tank3 Valve Error', class Errors, trigger "ALARMS" bit 14
   10: 'Tank3 Level L', class Warnings, trigger "ALARMS" bit 9

screen "Overview" 1280x800
   DateTimeField "Date/time field_1" at 1062,14 size 206x25
   TextField "Text field_1" at 241,471 size 117x44; Text 'Tank 1'
   TextField "Text field_2" at 569,474 size 117x44; Text 'Tank 2'
   TextField "Text field_3" at 883,474 size 117x44; Text 'Tank 3'
   SymbolLibrary "Symbol library_2" at 175,132 size 232x322
      ProcessValue <- "T1_LVL"
   Bar "Bar_4" at 176,144 size 230x292; Unit cm; MinimumValue 0; MaximumValue 300
      ProcessValue <- "T1_LVL"
   SymbolLibrary "Symbol library_1" at 507,138 size 232x322
   Bar "Bar_1" at 508,150 size 230x292; Unit cm; MinimumValue 0; MaximumValue 300
      ProcessValue <- "T2_LVL"
   SymbolLibrary "Symbol library_3" at 826,138 size 232x322
   Bar "Bar_2" at 827,150 size 230x292; Unit cm; MinimumValue 0; MaximumValue 300
      ProcessValue <- "T3_LVL"
   Button "Button_1" at 173,108 size 236x353; TextOff 'Text'
      on Press: ActivateScreen("Tank 1", 0)
   Button "Button_2" at 504,126 size 236x344; TextOff 'Text'
      on Press: ActivateScreen("Tank 2", 0)
   Button "Button_3" at 827,118 size 232x355; TextOff 'Text'
      on Press: ActivateScreen("Tank 3", 0)
   Button "Button_4" at 1100,708 size 139x64; TextOff 'ALARMS'
      on Press: ActivateScreen("Alarms", 0)

screen "Tank 1" 1280x800
   SymbolLibrary "Symbol library_2" at 151,101 size 232x322
   SymbolLibrary "Symbol library_3" at 404,336 size 89x73
   SymbolLibrary "Symbol library_4" at 515,355 size 70x52
   Bar "Bar_1" at 152,113 size 230x292; Unit cm; MinimumValue 0; MaximumValue 300
      ProcessValue <- "T1_LVL"
   SymbolLibrary "Symbol library_1" at 37,69 size 89x73
   TrendView "Trend view_1" at 626,116 size 600x300
   IOField "I/O field_1" at 411,291 size 81x32; FormatPattern 999; Unit  %
      ProcessValue <- "T1_Dis"
   IOField "I/O field_2" at 514,418 size 81x32; FormatPattern 999; Unit  %
      ProcessValue <- "T1_Dis_fl"
   IOField "I/O field_3" at 51,24 size 81x32; FormatPattern 999; Unit  %
      ProcessValue <- "T1_MV"
   TextField "Text field_1" at 821,478 size 226x33; Text 'CONTROL SYSTEM'
   Button "Button_1" at 51,732 size 104x40; TextOff 'MAIN'
      on Press: ActivateScreen("Overview", 0)
   DateTimeField "Date/time field_1" at 1062,14 size 206x25
   TextField "Text field_2" at 714,555 size 77x22; Text 'Setpoint:'
   TextField "Text field_3" at 714,615 size 94x22; Text 'Hysteresis:'
   IOField "I/O field_4" at 842,547 size 96x32; FormatPattern 999; Unit  cm
      ProcessValue <- "T1_SP"
   IOField "I/O field_5" at 843,609 size 96x32; FormatPattern 99.9; Unit  cm
      ProcessValue <- "T1_H_reg"
   IOField "I/O field_6" at 842,676 size 96x32; FormatPattern 999.9; Unit  %
      ProcessValue <- "T1_B_reg"
   TextField "Text field_4" at 714,678 size 95x22; Text 'Relay Gain:'

screen "Tank 2" 1280x800
   SymbolLibrary "Symbol library_2" at 151,101 size 232x322
   SymbolLibrary "Symbol library_3" at 404,336 size 89x73
   SymbolLibrary "Symbol library_4" at 515,355 size 70x52
   Bar "Bar_1" at 152,113 size 230x292; Unit cm; MinimumValue 0; MaximumValue 300
      ProcessValue <- "T2_LVL"
   SymbolLibrary "Symbol library_1" at 37,69 size 89x73
   TrendView "Trend view_1" at 626,116 size 600x328
   IOField "I/O field_1" at 411,291 size 81x32; FormatPattern 999; Unit  %
      ProcessValue <- "T2_Dis"
   IOField "I/O field_2" at 514,418 size 81x32; FormatPattern 999; Unit  %
      ProcessValue <- "T2_Dis_fl"
   IOField "I/O field_3" at 51,24 size 81x32; FormatPattern 999; Unit  %
      ProcessValue <- "T2_MV"
   TextField "Text field_1" at 821,478 size 226x33; Text 'CONTROL SYSTEM'
   Button "Button_1" at 51,732 size 104x40; TextOff 'MAIN'
      on Press: ActivateScreen("Overview", 0)
   DateTimeField "Date/time field_1" at 1062,14 size 206x25
   TextField "Text field_2" at 714,555 size 77x22; Text 'Setpoint:'
   TextField "Text field_3" at 714,612 size 67x22; Text 'Gain (P)'
   IOField "I/O field_4" at 867,547 size 96x32; FormatPattern 999; Unit  cm
      ProcessValue <- "T2_SP"
   IOField "I/O field_5" at 868,609 size 96x32; FormatPattern 999
      ProcessValue <- "T2_P_reg"
   IOField "I/O field_6" at 867,676 size 96x32; FormatPattern 999.9; Unit  s
      ProcessValue <- "T2_I_reg"
   TextField "Text field_4" at 714,678 size 138x22; Text 'Integral Time (Ti)'

screen "Tank 3" 1280x800
   TrendView "Trend view_1" at 626,116 size 600x328
   TextField "Text field_1" at 821,478 size 226x33; Text 'CONTROL SYSTEM'
   Button "Button_1" at 51,732 size 104x40; TextOff 'MAIN'
      on Press: ActivateScreen("Overview", 0)
   DateTimeField "Date/time field_1" at 1062,14 size 206x25
   SymbolLibrary "Symbol library_2" at 151,101 size 232x322
   SymbolLibrary "Symbol library_3" at 404,336 size 89x73
   SymbolLibrary "Symbol library_4" at 515,355 size 70x52
   Bar "Bar_1" at 152,113 size 230x292; Unit cm; MinimumValue 0; MaximumValue 300
      ProcessValue <- "T2_LVL"
   SymbolLibrary "Symbol library_1" at 37,69 size 89x73
   IOField "I/O field_1" at 411,291 size 81x32; FormatPattern 999; Unit  %
      ProcessValue <- "T3_Dis"
   IOField "I/O field_2" at 514,418 size 81x32; FormatPattern 999; Unit  %
      ProcessValue <- "T3_Dis_fl"
   IOField "I/O field_3" at 51,24 size 81x32; FormatPattern 999; Unit  %
      ProcessValue <- "T3_MV"
   TextField "Text field_2" at 674,571 size 77x22; Text 'Setpoint:'
   TextField "Text field_3" at 958,568 size 67x22; Text 'Gain (P)'
   IOField "I/O field_4" at 787,563 size 96x32; FormatPattern 999; Unit  cm
      ProcessValue <- "T3_SP"
   IOField "I/O field_5" at 1112,565 size 96x32; FormatPattern 999
      ProcessValue <- "T3_P_reg"
   IOField "I/O field_6" at 1111,632 size 96x32; FormatPattern 999.9; Unit  s
      ProcessValue <- "T3_I_reg"
   TextField "Text field_4" at 958,634 size 138x22; Text 'Integral Time (Ti)'
   IOField "I/O field_7" at 787,634 size 96x32; FormatPattern 999.9; Unit  %
      ProcessValue <- "T3_B_reg"
   TextField "Text field_5" at 674,638 size 93x22; Text 'Relay gain:'

screen "Alarms" 1280x800
   Button "Button_1" at 51,732 size 104x40; TextOff 'MAIN'
      on Press: ActivateScreen("Overview", 0)
   AlarmView "Alarm view_1" at 115,58 size 1065x549
   DateTimeField "Date/time field_1" at 1062,14 size 206x25
   Button "Button_2" at 292,622 size 182x76; TextOff 'Ackonowledge Tank 1'
      on Press: function_b14e0dd5("Acknowledge", 0); function_b14e0dd5("Acknowledge", 3); function_b14e0dd5("Acknowledge", 12)
   Button "Button_3" at 518,622 size 182x76; TextOff 'Ackonowledge Tank 2'
      on Press: function_b14e0dd5("Acknowledge", 4); function_b14e0dd5("Acknowledge", 7); function_b14e0dd5("Acknowledge", 13)
   Button "Button_4" at 735,620 size 182x76; TextOff 'Ackonowledge Tank 3'
      on Press: function_b14e0dd5("Acknowledge", 8); function_b14e0dd5("Acknowledge", 11); function_b14e0dd5("Acknowledge", 14)
   Button "Button_5" at 1000,620 size 182x76; TextOff 'Clear all'
      on Press: function_e14cd482(0)
*)

(* ===== HMI "HMI_RT_1" =====

ScreenModuleEditorView "Faceplate_1" 640x480
   Button "Button_1" at 10,10 size 96x32; TextOff 'Text'
*)

(* ===== HMI "HMI_RT_1" =====

ScreenModuleEditorView "Faceplate_1" 640x480
   Button "Button_1" at 10,10 size 96x32; TextOff 'Text'
*)